(* Logix 5000 project; controller NWGG 1756-L72 rev 35.12; software revision 35.00; part 9 of 19 *)
(* tags used below, declared in another part *)
   _25_16_1 : ALIAS FOR N200[11];
   _25_16_2 : ALIAS FOR N200[12];
   _25_16_3 : ALIAS FOR N200[13];
   _700_PROBE : ALIAS FOR T22[9];
   _700_TREAT : ALIAS FOR I7.3;
   _701K_GATE : ALIAS FOR B21[11].0;
   _701K_GATE1 : ALIAS FOR B21[11].1;
   _701K_GATE2 : ALIAS FOR B21[11].2;
   _708_BOT_CN : ALIAS FOR C5[5];
   _708G_BIN_1 : ALIAS FOR O9.15;
   _708G_BIN_2 : ALIAS FOR I7.4;
   _708G_CB13 : ALIAS FOR B21[8].0;
   _708G_CB131 : ALIAS FOR B21[8].1;
   _708G_CB132 : ALIAS FOR B21[8].2;
   _708G_HOLD : ALIAS FOR B21[8].3;
   _708G_HOLD1 : ALIAS FOR B21[8].6;
   _708G_RELEA : ALIAS FOR B21[8].4;
   _708G_RESET : ALIAS FOR B21[8].5;
   _709_BOT_CN : ALIAS FOR C5[6];
   _709G_BIN_1 : ALIAS FOR O10.15;
   _709G_BIN_2 : ALIAS FOR I7.5;
   _709G_CB19 : ALIAS FOR B21[9].0;
   _709G_CB191 : ALIAS FOR B21[9].1;
   _709G_CB192 : ALIAS FOR B21[9].2;
   _709G_HOLD : ALIAS FOR B21[9].3;
   _709G_HOLD1 : ALIAS FOR B21[9].6;
   _709G_RELEA : ALIAS FOR B21[9].4;
   _709G_RESET : ALIAS FOR B21[9].5;
   _709G_RUN_T : ALIAS FOR T22[8];
   _709G_TREAT : ALIAS FOR B21[9].7;
   _709G_TREAT1 : ALIAS FOR T22[10];
   A18 : INT[100];
   A_HOLD_MB : ALIAS FOR B3[1].3;
   A_TREATER : ALIAS FOR I24[6].8;
   B3 : DINT[250];
   Beta : BOOL;
   BIN_1_CLOSE : BOOL;
   BIN_1_OPEN : BOOL;
   BIN_2_CLOSE : BOOL;
   BIN_2_OPEN : BOOL;
   BIN_3_CLOSE : BOOL;
   BIN_3_OPEN : BOOL;
   BIN_4_CLOSE : BOOL;
   BIN_4_OPEN : BOOL;
   BIN_5_CLOSE : BOOL;
   BIN_5_OPEN : BOOL;
   BIN_6_CLOSE : BOOL;
   BIN_6_OPEN : BOOL;
   BIN_7_CLOSE : BOOL;
   BIN_7_OPEN : BOOL;
   CONC13_OP : ALIAS FOR A18[3];
   CONC13_SET : ALIAS FOR A18[0];
   CONC13_SET1 : ALIAS FOR B21[8].14;
   CONC19_OP : ALIAS FOR A18[13];
   CONC19_SET : ALIAS FOR B21[9].14;
   CONC_13_NO : ALIAS FOR B21[8].15;
   CONC_19_NO : ALIAS FOR B21[9].15;
   CONC_19_SE : ALIAS FOR A18[10];
   I24_006_Bit02 : ALIAS FOR I24[6].2;
   MAIN_TIMER1 : ALIAS FOR T11[1];
   N24 : DINT[31];
   N27 : DINT[50];
   N28 : DINT[17];
   N7 : DINT[100];
   O24 : INT[32];
   O24_007_Bit11 : ALIAS FOR O24[7].11;
   O24_007_Bit12 : ALIAS FOR O24[7].12;
   O24_007_Bit14 : ALIAS FOR O24[7].14;
   O25_012_Bit01 : ALIAS FOR O25[12].1;
   O25_012_Bit02 : ALIAS FOR O25[12].2;
   O25_012_Bit03 : ALIAS FOR O25[12].3;
   O25_012_Bit04 : ALIAS FOR O25[12].4;
   O25_012_Bit05 : ALIAS FOR O25[12].5;
   O25_012_Bit06 : ALIAS FOR O25[12].6;
   O25_012_Bit07 : ALIAS FOR O25[12].7;
   O25_012_Bit08 : ALIAS FOR O25[12].8;
   O25_012_Bit09 : ALIAS FOR O25[12].9;
   O25_012_Bit10 : ALIAS FOR O25[12].10;
   O25_012_Bit11 : ALIAS FOR O25[12].11;
   O25_012_Bit12 : ALIAS FOR O25[12].12;
   O25_012_Bit13 : ALIAS FOR O25[12].13;
   O25_012_Bit14 : ALIAS FOR O25[12].14;
   P_RESET_AU : ALIAS FOR B3[4].0;
   PMP_15_OFF_DLY : REAL;
   PMP_15_OFF_DLY_SCALE : REAL;
   PMP_15_ON_DLY : REAL;
   PMP_15_ON_DLY_SCALE : REAL;
   PMP_15_TMR : TIMER;
   PMP_15_TMR_2 : TIMER;
   PUMP_15_AUTO : BOOL;
   SCP_AOI : SCP_Inv[8];
   T11_TREAT : ALIAS FOR B3[11].0;
   T12_TREAT : ALIAS FOR B3[12].0;
   T13_TREAT : ALIAS FOR B3[13].0;
   T14_TREAT : ALIAS FOR B3[14].0;
   T15_TREAT : ALIAS FOR B3[15].0;
   T16_TREAT : ALIAS FOR B3[16].0;
   T17_TREAT : ALIAS FOR B3[17].0;
   T21_TREAT : ALIAS FOR B3[21].0;
   T22_TREAT : ALIAS FOR B3[22].0;
   T23_TREAT : ALIAS FOR B3[23].0;
   T24_TREAT : ALIAS FOR B3[24].0;
   T25 : TIMER[9];
   T25_TREAT : ALIAS FOR B3[25].0;
   T26_TREAT : ALIAS FOR B3[26].0;
   T27_TREAT : ALIAS FOR B3[27].0;
   T28_TREAT : ALIAS FOR B3[28].0;
   T29_TREAT : ALIAS FOR B3[29].0;
(* _2_MAIN, continued *)

ROUTINE _42_CONC_GATES   (* ladder *)
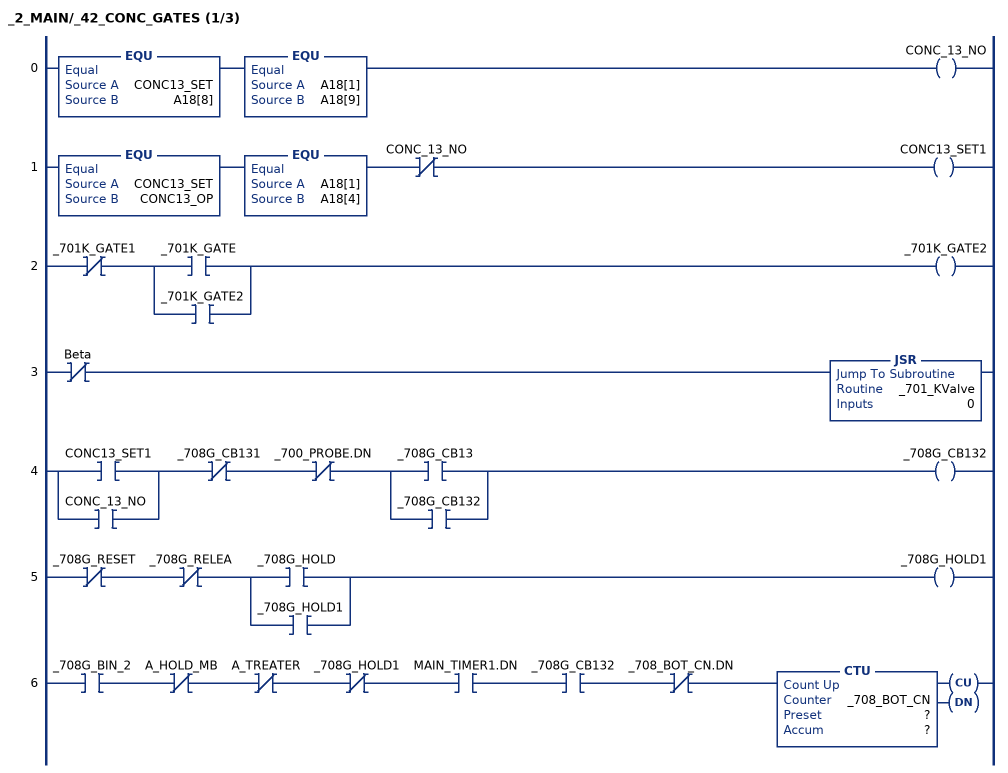
   0: EQU(CONC13_SET,A18[8])EQU(A18[1],A18[9])OTE(CONC_13_NO);
   1: EQU(CONC13_SET,CONC13_OP)EQU(A18[1],A18[4])XIO(CONC_13_NO)OTE(CONC13_SET1);
   2: XIO(_701K_GATE1)[XIC(_701K_GATE) ,XIC(_701K_GATE2) ]OTE(_701K_GATE2);
   3: XIO(Beta)JSR(_701_KValve,0);
   4: [XIC(CONC13_SET1) ,XIC(CONC_13_NO) ]XIO(_708G_CB131)XIO(_700_PROBE.DN)[XIC(_708G_CB13) ,XIC(_708G_CB132) ]OTE(_708G_CB132);
   5: XIO(_708G_RESET)XIO(_708G_RELEA)[XIC(_708G_HOLD) ,XIC(_708G_HOLD1) ]OTE(_708G_HOLD1);
   6: XIC(_708G_BIN_2)XIO(A_HOLD_MB)XIO(A_TREATER)XIO(_708G_HOLD1)XIC(MAIN_TIMER1.DN)XIC(_708G_CB132)XIO(_708_BOT_CN.DN)CTU(_708_BOT_CN,?,?);
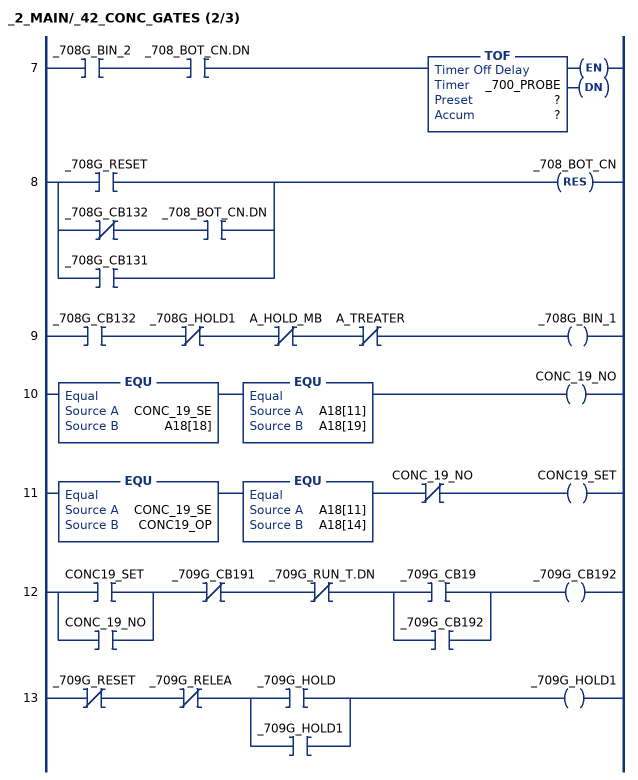
   7: XIC(_708G_BIN_2)XIC(_708_BOT_CN.DN)TOF(_700_PROBE,?,?);
   8: [XIC(_708G_RESET) ,XIO(_708G_CB132) XIC(_708_BOT_CN.DN) ,XIC(_708G_CB131) ]RES(_708_BOT_CN);
   9: XIC(_708G_CB132)XIO(_708G_HOLD1)XIO(A_HOLD_MB)XIO(A_TREATER)OTE(_708G_BIN_1);
   10: EQU(CONC_19_SE,A18[18])EQU(A18[11],A18[19])OTE(CONC_19_NO);
   11: EQU(CONC_19_SE,CONC19_OP)EQU(A18[11],A18[14])XIO(CONC_19_NO)OTE(CONC19_SET);
   12: [XIC(CONC19_SET) ,XIC(CONC_19_NO) ]XIO(_709G_CB191)XIO(_709G_RUN_T.DN)[XIC(_709G_CB19) ,XIC(_709G_CB192) ]OTE(_709G_CB192);
   13: XIO(_709G_RESET)XIO(_709G_RELEA)[XIC(_709G_HOLD) ,XIC(_709G_HOLD1) ]OTE(_709G_HOLD1);
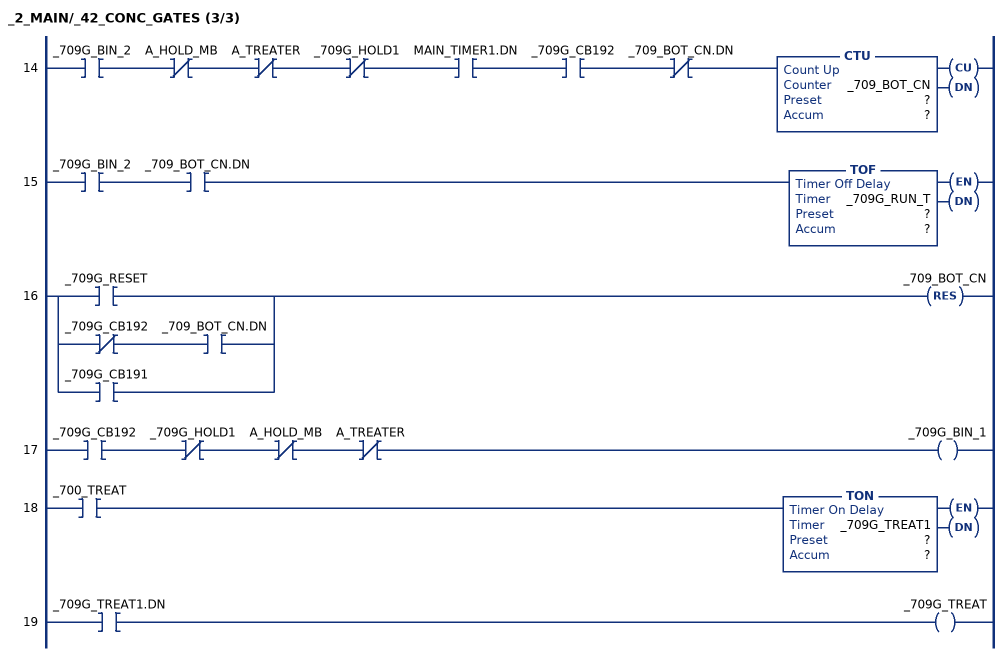
   14: XIC(_709G_BIN_2)XIO(A_HOLD_MB)XIO(A_TREATER)XIO(_709G_HOLD1)XIC(MAIN_TIMER1.DN)XIC(_709G_CB192)XIO(_709_BOT_CN.DN)CTU(_709_BOT_CN,?,?);
   15: XIC(_709G_BIN_2)XIC(_709_BOT_CN.DN)TOF(_709G_RUN_T,?,?);
   16: [XIC(_709G_RESET) ,XIO(_709G_CB192) XIC(_709_BOT_CN.DN) ,XIC(_709G_CB191) ]RES(_709_BOT_CN);
   17: XIC(_709G_CB192)XIO(_709G_HOLD1)XIO(A_HOLD_MB)XIO(A_TREATER)OTE(_709G_BIN_1);
   18: XIC(_700_TREAT)TON(_709G_TREAT1,?,?);
   19: XIC(_709G_TREAT1.DN)OTE(_709G_TREAT);
END_ROUTINE

ROUTINE _43_25_19_IE8   (* ladder *)
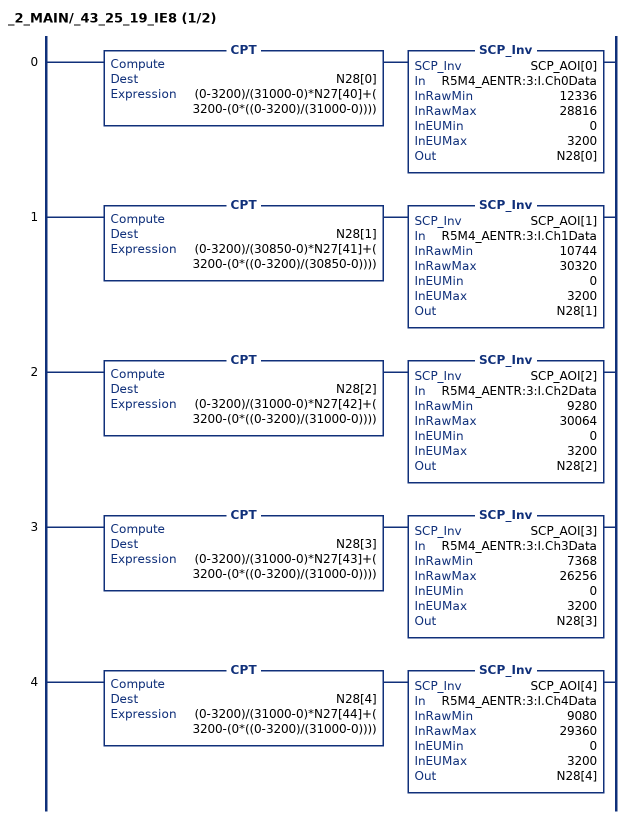
   0: CPT(N28[0],(0-3200)/(31000-0)*N27[40]+(3200-(0*((0-3200)/(31000-0)))))SCP_Inv(SCP_AOI[0],R5M4_AENTR:3:I.Ch0Data,12336,28816,0,3200,N28[0]);
   1: CPT(N28[1],(0-3200)/(30850-0)*N27[41]+(3200-(0*((0-3200)/(30850-0)))))SCP_Inv(SCP_AOI[1],R5M4_AENTR:3:I.Ch1Data,10744,30320,0,3200,N28[1]);
   2: CPT(N28[2],(0-3200)/(31000-0)*N27[42]+(3200-(0*((0-3200)/(31000-0)))))SCP_Inv(SCP_AOI[2],R5M4_AENTR:3:I.Ch2Data,9280,30064,0,3200,N28[2]);
   3: CPT(N28[3],(0-3200)/(31000-0)*N27[43]+(3200-(0*((0-3200)/(31000-0)))))SCP_Inv(SCP_AOI[3],R5M4_AENTR:3:I.Ch3Data,7368,26256,0,3200,N28[3]);
   4: CPT(N28[4],(0-3200)/(31000-0)*N27[44]+(3200-(0*((0-3200)/(31000-0)))))SCP_Inv(SCP_AOI[4],R5M4_AENTR:3:I.Ch4Data,9080,29360,0,3200,N28[4]);
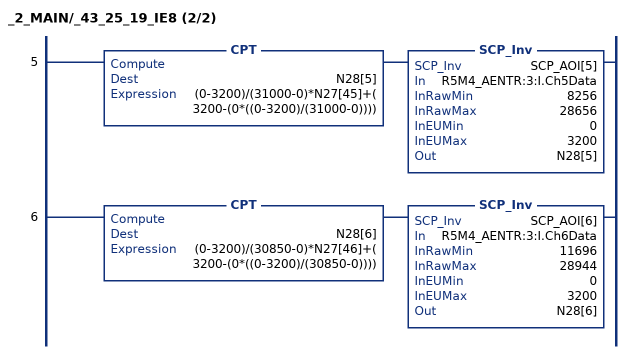
   5: CPT(N28[5],(0-3200)/(31000-0)*N27[45]+(3200-(0*((0-3200)/(31000-0)))))SCP_Inv(SCP_AOI[5],R5M4_AENTR:3:I.Ch5Data,8256,28656,0,3200,N28[5]);
   6: CPT(N28[6],(0-3200)/(30850-0)*N27[46]+(3200-(0*((0-3200)/(30850-0)))))SCP_Inv(SCP_AOI[6],R5M4_AENTR:3:I.Ch6Data,11696,28944,0,3200,N28[6]);
END_ROUTINE

ROUTINE _44_BINS_1_7   (* ladder *)
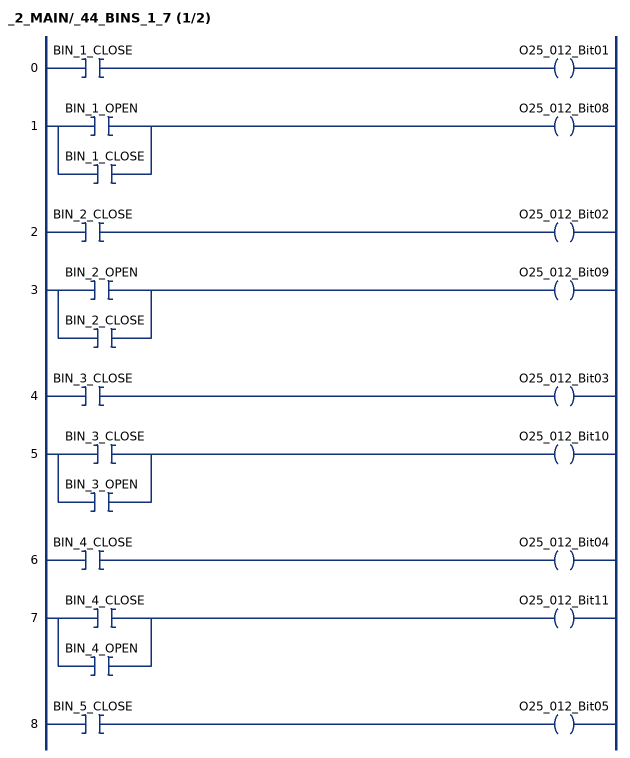
   0: XIC(BIN_1_CLOSE)OTE(O25_012_Bit01);
   1: [XIC(BIN_1_OPEN) ,XIC(BIN_1_CLOSE) ]OTE(O25_012_Bit08);
   2: XIC(BIN_2_CLOSE)OTE(O25_012_Bit02);
   3: [XIC(BIN_2_OPEN) ,XIC(BIN_2_CLOSE) ]OTE(O25_012_Bit09);
   4: XIC(BIN_3_CLOSE)OTE(O25_012_Bit03);
   5: [XIC(BIN_3_CLOSE) ,XIC(BIN_3_OPEN) ]OTE(O25_012_Bit10);
   6: XIC(BIN_4_CLOSE)OTE(O25_012_Bit04);
   7: [XIC(BIN_4_CLOSE) ,XIC(BIN_4_OPEN) ]OTE(O25_012_Bit11);
   8: XIC(BIN_5_CLOSE)OTE(O25_012_Bit05);
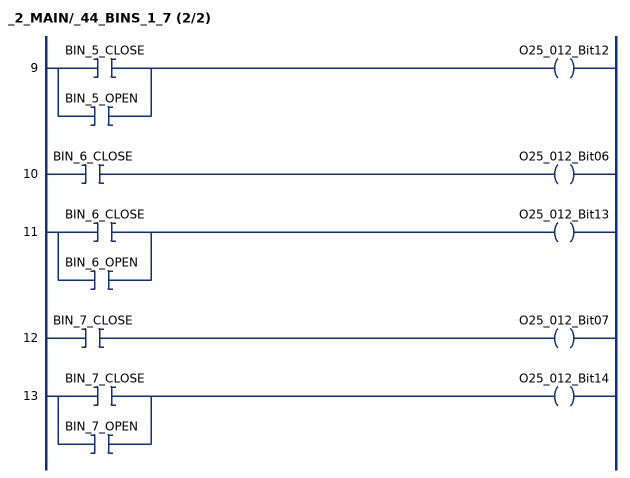
   9: [XIC(BIN_5_CLOSE) ,XIC(BIN_5_OPEN) ]OTE(O25_012_Bit12);
   10: XIC(BIN_6_CLOSE)OTE(O25_012_Bit06);
   11: [XIC(BIN_6_CLOSE) ,XIC(BIN_6_OPEN) ]OTE(O25_012_Bit13);
   12: XIC(BIN_7_CLOSE)OTE(O25_012_Bit07);
   13: [XIC(BIN_7_CLOSE) ,XIC(BIN_7_OPEN) ]OTE(O25_012_Bit14);
END_ROUTINE

ROUTINE _45_PMP_11_14   (* ladder *)
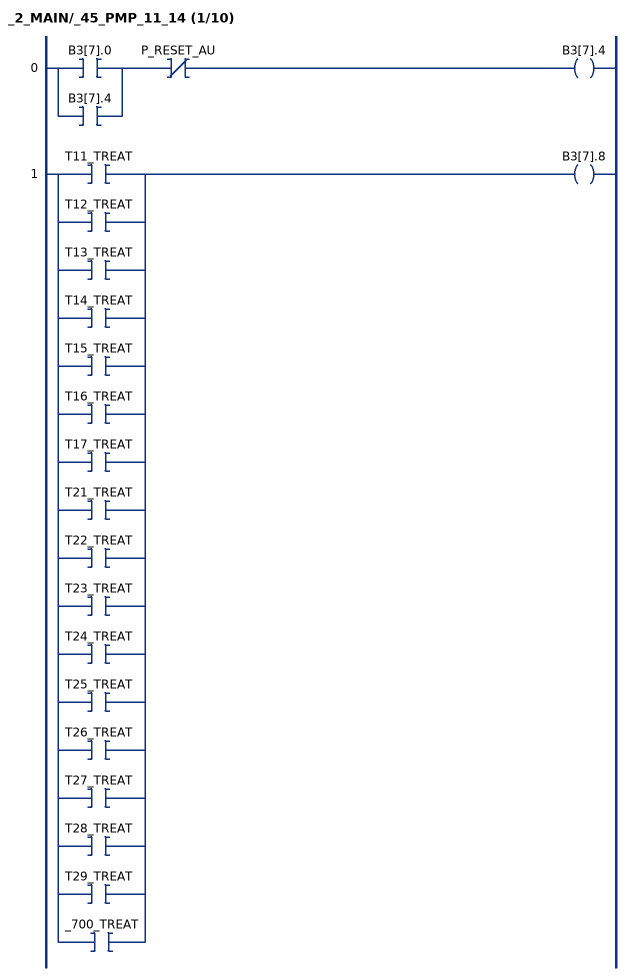
   0: [XIC(B3[7].0) ,XIC(B3[7].4) ]XIO(P_RESET_AU)OTE(B3[7].4);
   1: [XIC(T11_TREAT) ,XIC(T12_TREAT) ,XIC(T13_TREAT) ,XIC(T14_TREAT) ,XIC(T15_TREAT) ,XIC(T16_TREAT) ,XIC(T17_TREAT) ,XIC(T21_TREAT) ,XIC(T22_TREAT) ,XIC(T23_TREAT) ,XIC(T24_TREAT) ,XIC(T25_TREAT) ,XIC(T26_TREAT) ,XIC(T27_TREAT) ,XIC(T28_TREAT) ,XIC(T29_TREAT) ,XIC(_700_TREAT) ]OTE(B3[7].8);
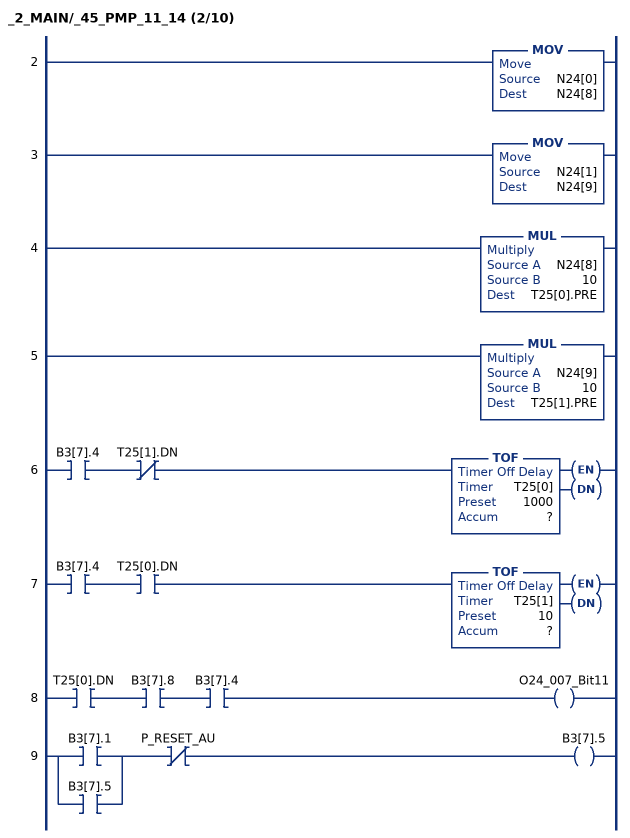
   2: MOV(N24[0],N24[8]);
   3: MOV(N24[1],N24[9]);
   4: MUL(N24[8],10,T25[0].PRE);
   5: MUL(N24[9],10,T25[1].PRE);
   6: XIC(B3[7].4)XIO(T25[1].DN)TOF(T25[0],?,?);
   7: XIC(B3[7].4)XIC(T25[0].DN)TOF(T25[1],?,?);
   8: XIC(T25[0].DN)XIC(B3[7].8)XIC(B3[7].4)OTE(O24_007_Bit11);
   9: [XIC(B3[7].1) ,XIC(B3[7].5) ]XIO(P_RESET_AU)OTE(B3[7].5);
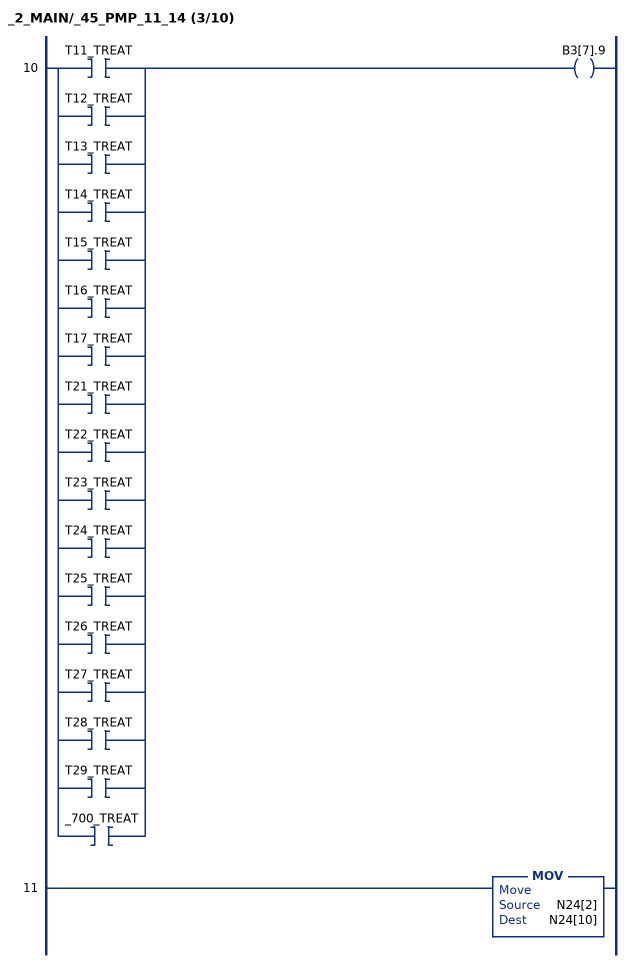
   10: [XIC(T11_TREAT) ,XIC(T12_TREAT) ,XIC(T13_TREAT) ,XIC(T14_TREAT) ,XIC(T15_TREAT) ,XIC(T16_TREAT) ,XIC(T17_TREAT) ,XIC(T21_TREAT) ,XIC(T22_TREAT) ,XIC(T23_TREAT) ,XIC(T24_TREAT) ,XIC(T25_TREAT) ,XIC(T26_TREAT) ,XIC(T27_TREAT) ,XIC(T28_TREAT) ,XIC(T29_TREAT) ,XIC(_700_TREAT) ]OTE(B3[7].9);
   11: MOV(N24[2],N24[10]);
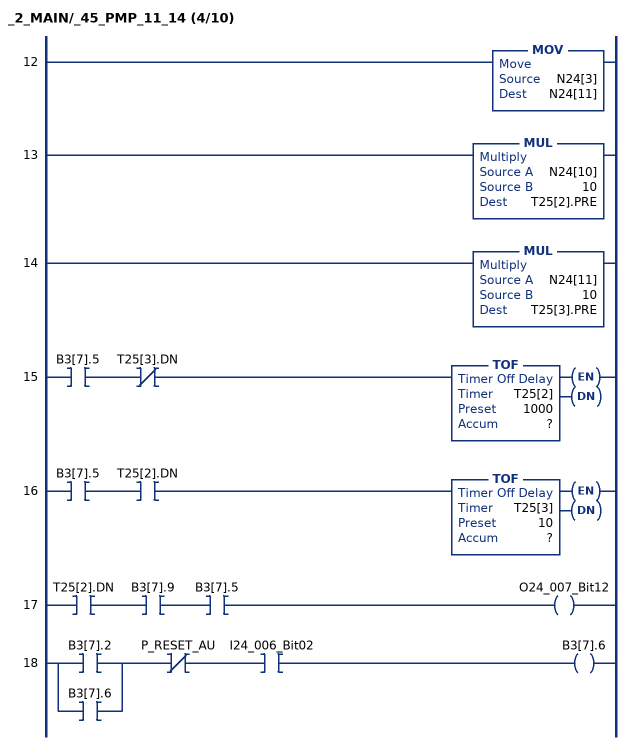
   12: MOV(N24[3],N24[11]);
   13: MUL(N24[10],10,T25[2].PRE);
   14: MUL(N24[11],10,T25[3].PRE);
   15: XIC(B3[7].5)XIO(T25[3].DN)TOF(T25[2],?,?);
   16: XIC(B3[7].5)XIC(T25[2].DN)TOF(T25[3],?,?);
   17: XIC(T25[2].DN)XIC(B3[7].9)XIC(B3[7].5)OTE(O24_007_Bit12);
   18: [XIC(B3[7].2) ,XIC(B3[7].6) ]XIO(P_RESET_AU)XIC(I24_006_Bit02)OTE(B3[7].6);
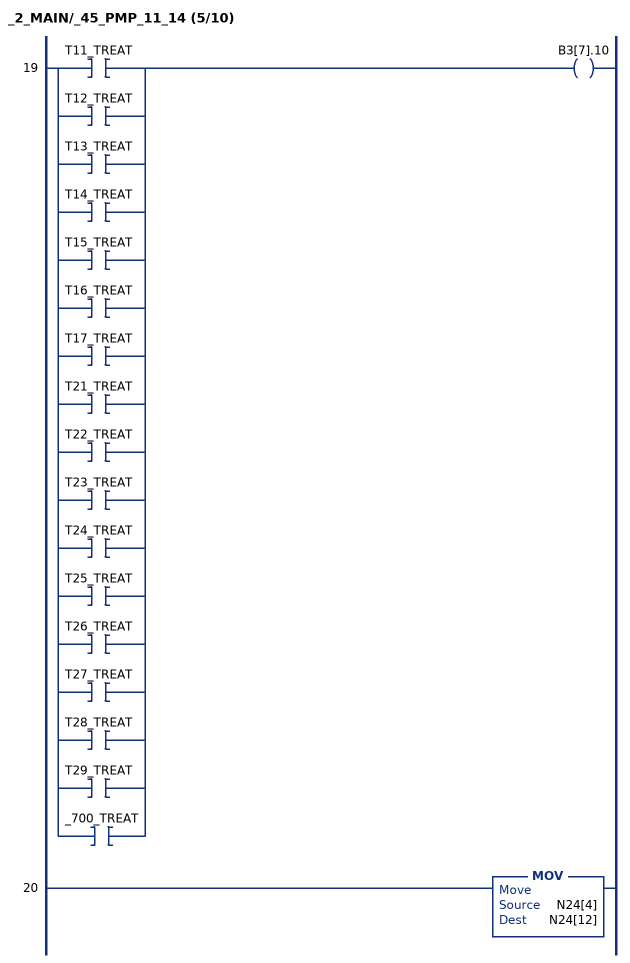
   19: [XIC(T11_TREAT) ,XIC(T12_TREAT) ,XIC(T13_TREAT) ,XIC(T14_TREAT) ,XIC(T15_TREAT) ,XIC(T16_TREAT) ,XIC(T17_TREAT) ,XIC(T21_TREAT) ,XIC(T22_TREAT) ,XIC(T23_TREAT) ,XIC(T24_TREAT) ,XIC(T25_TREAT) ,XIC(T26_TREAT) ,XIC(T27_TREAT) ,XIC(T28_TREAT) ,XIC(T29_TREAT) ,XIC(_700_TREAT) ]OTE(B3[7].10);
   20: MOV(N24[4],N24[12]);
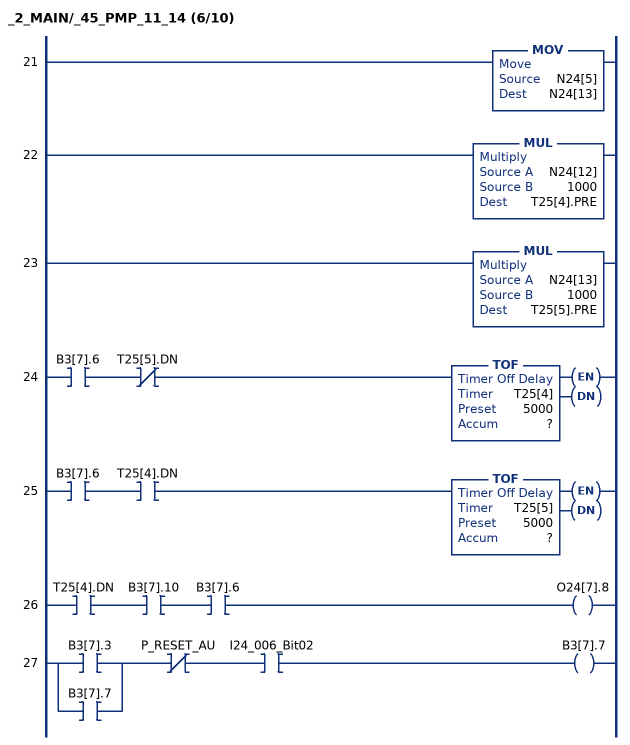
   21: MOV(N24[5],N24[13]);
   22: MUL(N24[12],1000,T25[4].PRE);
   23: MUL(N24[13],1000,T25[5].PRE);
   24: XIC(B3[7].6)XIO(T25[5].DN)TOF(T25[4],?,?);
   25: XIC(B3[7].6)XIC(T25[4].DN)TOF(T25[5],?,?);
   26: XIC(T25[4].DN)XIC(B3[7].10)XIC(B3[7].6)OTE(O24[7].8);
   27: [XIC(B3[7].3) ,XIC(B3[7].7) ]XIO(P_RESET_AU)XIC(I24_006_Bit02)OTE(B3[7].7);
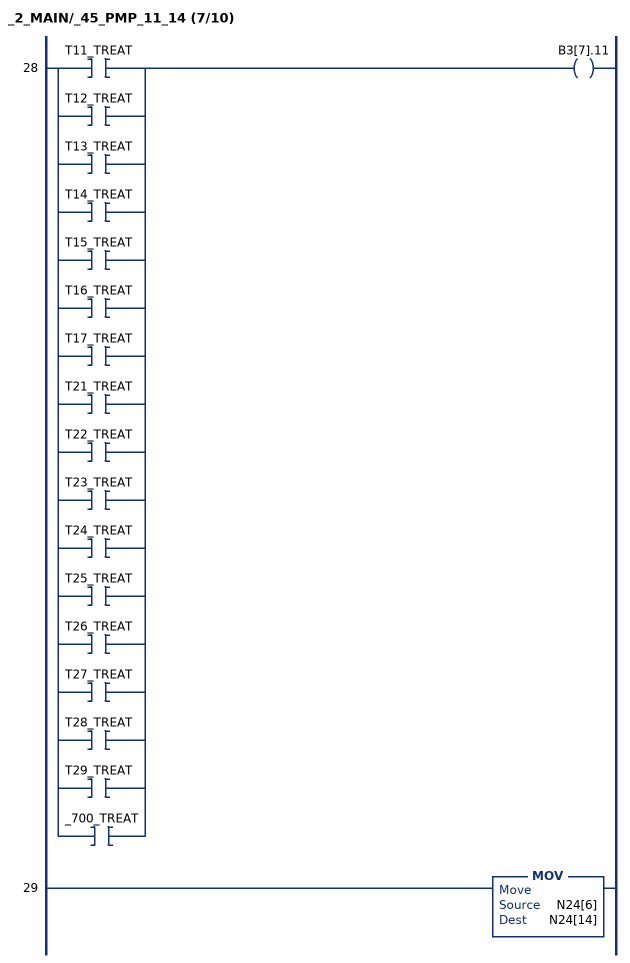
   28: [XIC(T11_TREAT) ,XIC(T12_TREAT) ,XIC(T13_TREAT) ,XIC(T14_TREAT) ,XIC(T15_TREAT) ,XIC(T16_TREAT) ,XIC(T17_TREAT) ,XIC(T21_TREAT) ,XIC(T22_TREAT) ,XIC(T23_TREAT) ,XIC(T24_TREAT) ,XIC(T25_TREAT) ,XIC(T26_TREAT) ,XIC(T27_TREAT) ,XIC(T28_TREAT) ,XIC(T29_TREAT) ,XIC(_700_TREAT) ]OTE(B3[7].11);
   29: MOV(N24[6],N24[14]);
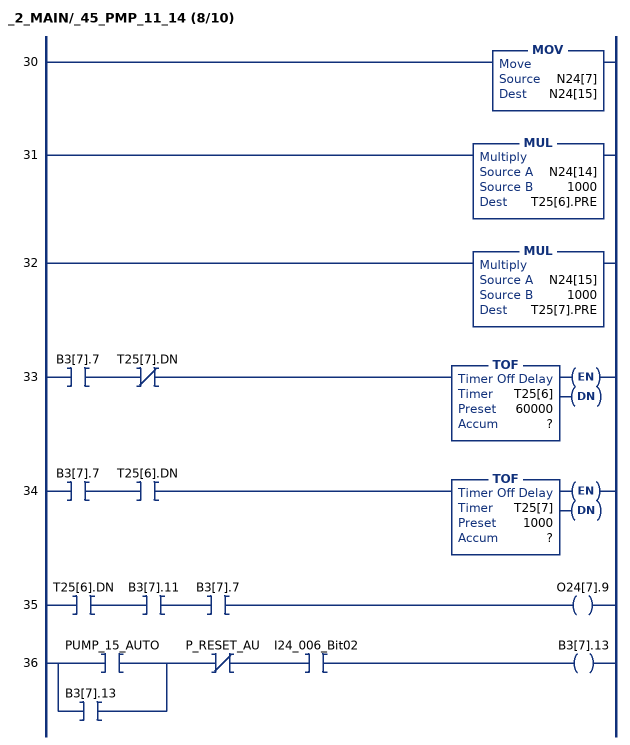
   30: MOV(N24[7],N24[15]);
   31: MUL(N24[14],1000,T25[6].PRE);
   32: MUL(N24[15],1000,T25[7].PRE);
   33: XIC(B3[7].7)XIO(T25[7].DN)TOF(T25[6],?,?);
   34: XIC(B3[7].7)XIC(T25[6].DN)TOF(T25[7],?,?);
   35: XIC(T25[6].DN)XIC(B3[7].11)XIC(B3[7].7)OTE(O24[7].9);
   36: [XIC(PUMP_15_AUTO) ,XIC(B3[7].13) ]XIO(P_RESET_AU)XIC(I24_006_Bit02)OTE(B3[7].13);
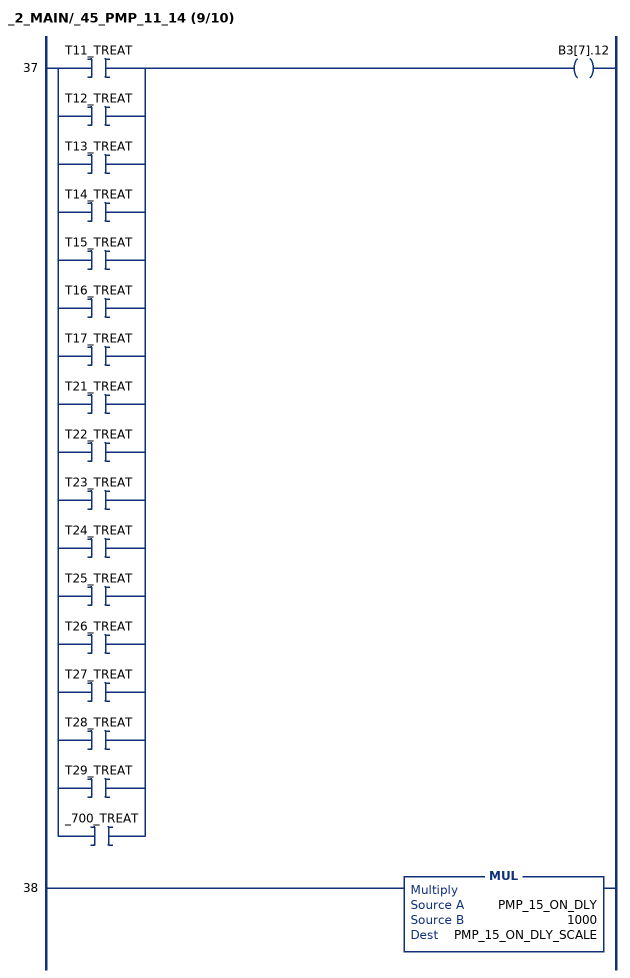
   37: [XIC(T11_TREAT) ,XIC(T12_TREAT) ,XIC(T13_TREAT) ,XIC(T14_TREAT) ,XIC(T15_TREAT) ,XIC(T16_TREAT) ,XIC(T17_TREAT) ,XIC(T21_TREAT) ,XIC(T22_TREAT) ,XIC(T23_TREAT) ,XIC(T24_TREAT) ,XIC(T25_TREAT) ,XIC(T26_TREAT) ,XIC(T27_TREAT) ,XIC(T28_TREAT) ,XIC(T29_TREAT) ,XIC(_700_TREAT) ]OTE(B3[7].12);
   38: MUL(PMP_15_ON_DLY,1000,PMP_15_ON_DLY_SCALE);
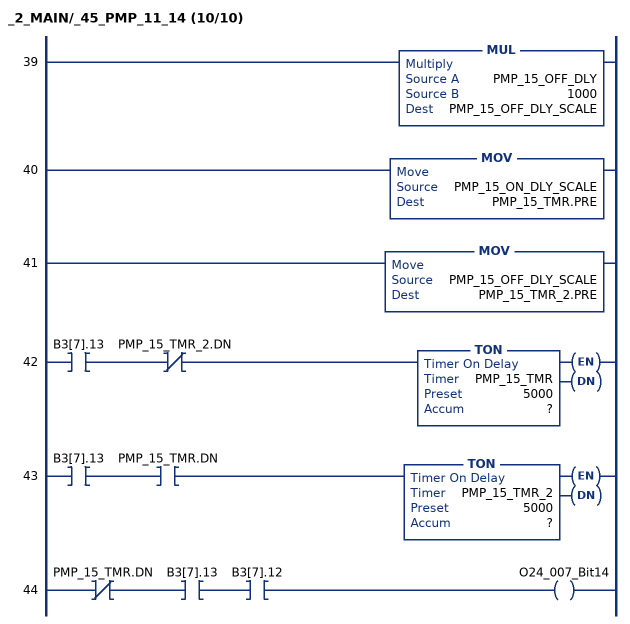
   39: MUL(PMP_15_OFF_DLY,1000,PMP_15_OFF_DLY_SCALE);
   40: MOV(PMP_15_ON_DLY_SCALE,PMP_15_TMR.PRE);
   41: MOV(PMP_15_OFF_DLY_SCALE,PMP_15_TMR_2.PRE);
   42: XIC(B3[7].13)XIO(PMP_15_TMR_2.DN)TON(PMP_15_TMR,?,?);
   43: XIC(B3[7].13)XIC(PMP_15_TMR.DN)TON(PMP_15_TMR_2,?,?);
   44: XIO(PMP_15_TMR.DN)XIC(B3[7].13)XIC(B3[7].12)OTE(O24_007_Bit14);
END_ROUTINE

ROUTINE _45_SCALING   (* function block diagram *)
   SHEET 1
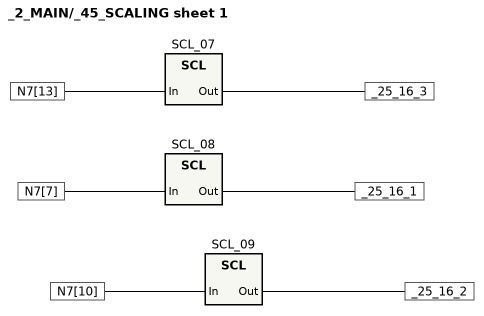
   SCL_07 : SCL(In := N7[13]);
   SCL_08 : SCL(In := N7[7]);
   SCL_09 : SCL(In := N7[10]);
   _25_16_1 := SCL_08.Out;
   _25_16_3 := SCL_07.Out;
   _25_16_2 := SCL_09.Out;
END_ROUTINE
